         A     "DB123_MH_IO_Signals".MH[1].IN.MH_Stop;
         A     "DB123_MH_IO_Signals".MH[1].IN.MH_Manual_Mode;
   //    O
   //    UN    "DB005_RS<->Extern".FT_01.Daten_von_FT.Schaeumvorbereitung
         O     "DB123_MH_IO_Signals".MH[1].IN.MH_Auto_Mode;
         =     #Stop_MH;

         A     "DB123_MH_IO_Signals".MH[1].IN.MH_Status.shotactive_MH;
         AN    "DB614_MH_State".InertingMH[1].Inert_ON_OFF;
         A     "DB619_State_MPart".ShotMa[1].ShotData.PurgeMH_AfterShot;
         A     "DB614_MH_State".MH_Status[1].Switch_Service_ON_OFF;
         S     "DB614_MH_State".InertingMH[1].Start_Prepare_Purge_after_Shot;

         A     "DB614_MH_State".InertingMH[1].Start_Prepare_Purge_after_Shot;
         A     "DB619_State_MPart".Cycle[1].PulsShotend;
         A     "IPS_CP_MH01";
         S     "DB614_MH_State".InertingMH[1].Start_Purge_after_Shot;

         AN    "IPS_CP_MH01";
   //      U(
   //      U     "DB614_MH_State".InertingMH[1].Reserve41
   //      O     "DB614_MH_State".InertingMH[1].Inert_ON_OFF
   //      )
         A     "DB704_MH_Value".MH_Inerting[1].with_Purge;
         S     "DB614_MH_State".InertingMH[1].Enable_Purge;

         A     "IPS_CP_MH01";
         A     "DB614_MH_State".InertingMH[1].Enable_Purge;
         FP    "DB614_MH_State".InertingMH[1].Reserve40;
         S     "DB614_MH_State".InertingMH[1].Reserve42;

         A     "T_CP_forward_MH01";
         A     "DB614_MH_State".InertingMH[1].Enable_Purge;
         AN    "DB619_State_MPart".Cycle[1].running;
         S     "DB614_MH_State".InertingMH[1].Start_Purge_Manual;

         A     "DB614_MH_State".InertingMH[1].Start_Purge_Manual;
         AN    "DB619_State_MPart".Cycle[1].running;
         AN    "IPS_CP_MH01";
         S     "DB614_MH_State".InertingMH[1].HF_Start_Purge_Manual;
         R     "DB614_MH_State".InertingMH[1].Start_Purge_Manual;

         A(;
         A     "DB614_MH_State".InertingMH[1].HF_Start_Purge_Manual;
         O     "DB614_MH_State".InertingMH[1].Reserve42;
         );
         A     "IPS_CP_MH01";
         L     "DB704_MH_Value".MH_Inerting[1].Purge_time;
         JC    BLAS;

         A     "DB614_MH_State".InertingMH[1].Start_Purge_after_Shot;
         L     "DB704_MH_Value".MH_Inerting[1].Purge_after_Shot;
   BLAS: SE    "TM_Purge_after_Shot";
         A     "TM_Purge_after_Shot";
         FN    "DB614_MH_State".InertingMH[1].FN_Purge_after_shot_finished;
         R     "DB614_MH_State".InertingMH[1].HF_Start_Purge_Manual;
         R     "DB614_MH_State".InertingMH[1].Start_Prepare_Purge_after_Shot;
         R     "DB614_MH_State".InertingMH[1].Start_Purge_after_Shot;
         R     "DB614_MH_State".InertingMH[1].Enable_Purge;
         R     "DB614_MH_State".InertingMH[1].Reserve42;

         A     "TM_Purge_after_Shot";
         =     #Purge_Manual;

         A     #Purge_Manual;
         A     "DB614_MH_State".InertingMH[1].Reserve41;
         L     S5T#1S;
         SD    "TM_Reset_after_purge";
         A     "TM_Reset_after_purge";
         R     "DB704_MH_Value".MH_Inerting[1].with_purge_after_Shot;
         R     "DB614_MH_State".InertingMH[1].Enable_Purge;
         R     "DB614_MH_State".InertingMH[1].Reserve42;
         R     "DB614_MH_State".InertingMH[1].Reserve41;
         R     "DB614_MH_State".InertingMH[1].Start_Prepare_Purge_after_Shot;
         R     "DB614_MH_State".InertingMH[1].Start_Purge_after_Shot;

         L     0.0;
         T     "DB704_MH_Value".MH_Inerting[1].Reference_Value_Inert;

   //      CALL  "FC118_Enable_Inerting"
   //         Prg_Number     :=#InertPRG
   //         Ps_Number      :=1      //"DB619_State_MPart".ToolMa[1].PartShot
   //         ReferenceValue :="DB704_MH_Value".MH_Inerting[1].Reference_Value_Inert
   //         Inerting_OFF   :="DB614_MH_State".InertingMH[1].Inert_ON_OFF
   //         Shotwight      :=#Shotwight
END_REGION

REGION Network 2: MH01: Valve Nitrogen for Inerting
         SET;
         =     "DB704_MH_Value".MH_Inerting[1].with_Cycle_before_Inert_finished;

         CALL  "FC116_Inerting"
         ( IN_Enable                        := "DB619_State_MPart".Cycle[1].Release,
           IN_With_Inerting                 := "DB704_MH_Value".Mixinghead[1].WithInerting,
           IN_OP_Mode_Manual                := "DB123_MH_IO_Signals".MH[1].IN.MH_Manual_Mode,
           IN_OP_Mode_Wetshot               := 1,  //"DB614_MH_State".MH_Status[1].Switch_Service_ON_OFF
           IN_OP_Mode_Test                  := "DB619_State_MPart".Operationmode[1].Test,
           IN_Start                         := #Start_MH,
           IN_Stop                          := #Stop_MH,
           IN_T_Flushing                    := FALSE,
           IN_T_Purge_Air                   := #Purge_Manual,
           IN_Enable_pressurize_time        := "DB704_MH_Value".MH_Inerting[1].with_Cycle_before_Inert_finished,
           IN_AutoPurge_Air                 := FALSE,
           IN_Quitt_Fault                   := "DB009_Faults".Faults_Reset_FKT_M1,
           IN_Cycle_runs                    := FALSE,
           IN_MC_Activ                      := "DB614_MH_State".MH_Status[1].Switch_Service_ON_OFF,
           IN_PressurizeTimeRuns            := "DB619_State_MPart".Cycle[1].PressurizeTimeRuns,
           IN_Shotend                       := "DB619_State_MPart".Cycle[1].LastShotinToolFinished,
           IN_S_P_N2                        := "P_Nitrogen_Inerting_OK",
           IN_S_P_FlushingAgent             := TRUE,
           IN_MH_selected                   := "DB619_State_MPart".SWU[1].SWU_released."01",
           IN_Inert_MH                      := "DB704_MH_Value".MH_Inerting[1].with_inert_over_MH,
           IN_Inert_Lance                   := "DB704_MH_Value".MH_Inerting[1].with_inert_over_Lance,
           IN_IntervalCleaning              := "DB704_MH_Value".MH_Inerting[1].with_Interval_Purge,
           IN_Ctrl_Fault_On                 := TRUE,
           IN_Flowrate_N2_Actual            := "DB614_MH_State".InertingMH[1].Actual_Flow_N2_Visu,
           IN_Shotwight                     := #Shotwight,
           IN_Foam_Density                  := "DB704_MH_Value".MH_Inerting[1].Foam_density,
           IN_Leakage_value                 := "DB704_MH_Value".MH_Inerting[1].Leakage_Value,
           IN_DW_P_Build_Up_Before_Shot     := "DB700_Machine".Machine[1].PressureBuildUpTime,
           IN_DW_MaxInertTime               := "DB704_MH_Value".MH_Inerting[1].Max_Inerting_Time,
           IN_DW_Delay_Purge                := "DB704_MH_Value".MH_Inerting[1].Delay_Purge,
           IN_DW_Ready_time                 := "DB704_MH_Value".MH_Inerting[1].Ready_Time_after_Inert,
           IN_DW_Purge_time                 := "DB704_MH_Value".MH_Inerting[1].Purge_time,
           IN_DW_Delay_Plunger              := "DB704_MH_Value".MH_Inerting[1].Delay_Plunger,
           IN_DW_Delay_IntervalCleaning     := "DB704_MH_Value".MH_Inerting[1].Delay_Purge_Interval,
           IN_DW_PurgeTime_IntervalCleaning := "DB704_MH_Value".MH_Inerting[1].Purge_Time_interval,
           IN_DW_PauseTime_IntervalCleaning := "DB704_MH_Value".MH_Inerting[1].Pause_Time_interval,
           IN_DW_Duration_IntervalCleaning  := "DB704_MH_Value".MH_Inerting[1].Duration_Time_Interval,
           IN_Timer_Delay_Leakage           := "T_Leakage_Ctrl_N2",
           IN_Timer_hourly_tact             := "T_Leakage_Ctrl_Tact_N2",
           IN_Timer_Inerting                := "T_Inerting",
           IN_Timer_Ready                   := "T_Ready_for_Shot",
           IN_Timer_Delay_Purge             := "T_Delay_Purge",
           IN_Timer_Purge                   := "T_Purge",
           IN_Timer_Maximum_InertTime       := "T_Max_Inerting",
           IN_Timer_Delay_Plunger_N2        := "T_Delay_Plunger",
           IN_Timer_Delay_Tact              := "T_Delay_Purge_Tact",
           IN_Timer_PurgeTime_Tact          := "T_Purge_Tact",
           IN_Timer_PauseTime_Tact          := "T_Pause_Tact",
           IN_Timer_TotalTime_Tact          := "T_Total_Time_Purge",
           OUT_H_Inert                      := #dummy,
           OUT_H_Purge                      := #dummy,
           OUT_H_FlushingAgent              := #dummy,
           IO_DD_Inertfactor                := "DB704_MH_Value".MH_Inerting[1].Inerting_factor,
           IO_DD_StartOffset                := "DB704_MH_Value".MH_Inerting[1].Start_Offset,
           IO_DD_DF_N2_SetValue             := "DB614_MH_State".InertingMH[1].Computed_Value,
           IO_DD_DF_N2_Total                := "DB614_MH_State".InertingMH[1].Total_Flow_N2_Visu,
           IO_DD_DF_N2_Leakage              := "DB614_MH_State".InertingMH[1].Leakage_Total_Flow_N2_Visu,
           IO_MH_Logged_on                  := #dummy,
           IO_V_Piston                      := "V_Inert_Piston_MH1",
           IO_V_Inert                       := #Inerting,
           IO_V_Purge_Air                   := #Purge,
           IO_V_FlushingAgent               := #dummy,
           IO_Status                        := "DB614_MH_State".InertingMH[1],
           IO_Status_Faults                 := "DB824_Error_MH_CP".InertingBlowOut_MH[1],
           IO_NewFault                      := "DB009_Faults".Faultschanging_M1,
           IO_FaultLevel_1                  := "DB009_Faults".Faults_FKT_Grp_1_M1,
           IO_FaultLevel_2                  := "DB009_Faults".Faults_FKT_Grp_2_M1,
           IO_FaultLevel_3                  := "DB009_Faults".Faults_FKT_Grp_3_M1
         );

         A     #Purge;
         O     #Inerting;
         =     "V_Inert_MH1";
END_REGION
END_FUNCTION_BLOCK

FUNCTION_BLOCK "FB120_ProcanIO_RW"   // FB120, STL
TITLE = Transfer IO-Values from and to the ProCan-Moduls
{ S7_Optimized_Access := 'FALSE' }
AUTHOR : KT242
NAME : StPUCSPS
VERSION : 0.1
   VAR_TEMP
      Temp_ShotTimeAct : Real;
      dummy : Bool;
      Null : Word;
      ERROR_CODE : Int;
   END_VAR
BEGIN

REGION Network 1: Reset adresses od flow and MH
END_REGION

REGION Network 2: Read input values of procan modul
   //
         CALL  "FC120_read_ProCan";
END_REGION

REGION Network 3: PV Shot time
         L     0;
         T     #Temp_ShotTimeAct;

         AN    "DB619_State_MPart".SWU[1].Open_SWU_allone."01";
         JC    szm2;
         L     "DB123_MH_IO_Signals".MH[1].IN.Shottime;
         JU    szpv;
   szm2: AN    "DB619_State_MPart".SWU[1].Open_SWU_allone."02";
         JC    szm3;
         L     "DB123_MH_IO_Signals".MH[2].IN.Shottime;
         JU    szpv;
   szm3: AN    "DB619_State_MPart".SWU[1].Open_SWU_allone."03";
         JC    szm4;
         L     "DB123_MH_IO_Signals".MH[3].IN.Shottime;
         JU    szpv;
   szm4: AN    "DB619_State_MPart".SWU[1].Open_SWU_allone."04";
         JC    szm5;
         L     "DB123_MH_IO_Signals".MH[4].IN.Shottime;
         JU    szpv;
   szm5: AN    "DB619_State_MPart".SWU[1].Open_SWU_allone."05";
         JC    szm6;
         L     "DB123_MH_IO_Signals".MH[5].IN.Shottime;
         JU    szpv;
   szm6: AN    "DB619_State_MPart".SWU[1].Open_SWU_allone."06";
         JC    szm7;
         L     "DB123_MH_IO_Signals".MH[6].IN.Shottime;
         JU    szpv;
   szm7: AN    "DB619_State_MPart".SWU[1].Open_SWU_allone."07";
         JC    szm8;
         L     "DB123_MH_IO_Signals".MH[7].IN.Shottime;
         JU    szpv;
   szm8: AN    "DB619_State_MPart".SWU[1].Open_SWU_allone."08";
         JC    szm9;
         L     "DB123_MH_IO_Signals".MH[8].IN.Shottime;
         JU    szpv;
   szm9: AN    "DB619_State_MPart".SWU[1].Open_SWU_allone."09";
         JC    szm10;
         L     "DB123_MH_IO_Signals".MH[9].IN.Shottime;
         JU    szpv;
   szm10:AN    "DB619_State_MPart".SWU[1].Open_SWU_allone."10";
         JC    szm11;
         L     "DB123_MH_IO_Signals".MH[10].IN.Shottime;
         JU    szpv;
   szm11:AN    "DB619_State_MPart".SWU[1].Open_SWU_allone."11";
         JC    szm12;
         L     "DB123_MH_IO_Signals".MH[11].IN.Shottime;
         JU    szpv;
   szm12:AN    "DB619_State_MPart".SWU[1].Open_SWU_allone."12";
         JC    szm13;
         L     "DB123_MH_IO_Signals".MH[12].IN.Shottime;
         JU    szpv;
   szm13:JU    send;

   szpv: T     #Temp_ShotTimeAct;

         CALL  "FC920_PV_Calc_Act_Value"
         ( IN_Act_Value_read := TRUE,
           IN_Act_Value_ext  := TRUE,
           IN_Ext_Value      := #Temp_ShotTimeAct,
           IN_Read_Double    := TRUE,
           IN_FLT_Needful    := TRUE,
           IN_FLT_Reset      := "DB009_Faults".Faults_Reset_FKT_M1,
           IO_Any_ArrayPV    := "DB606_PV_Machine".Machine[1].ShotTime,
           IO_Fault_Sensor   := #dummy,
           IO_New_Fault      := #dummy,
           IO_FLT_Level_3    := #dummy
         );

   send: NOP   0;
END_REGION

REGION Network 4: Write output values of procan modul
   // Ein beschreiben der Module für die Mischköpfe ist nur bei LFI- Mischköpfen oder 
   // bei weiteren Mischköopfen bei dennen der Durchfluß eines Mediums am Mischkopf 
   // aufgenommen und geregelt wird (z.B. Faser) nötig.
   //
         CALL  "FC126_write_ProCan";
END_REGION
END_FUNCTION_BLOCK

FUNCTION_BLOCK "FB916_PV_LimitControl"   // FB916, STL
TITLE = Read prozess values and limit control of process values
{ S7_Optimized_Access := 'FALSE' }
AUTHOR : KT242
VERSION : 0.1
   VAR_TEMP
      DInt_dummy : DInt;
      FLT_quit_from_PLC : Bool;
      NewFault : Bool;
      ErrorLevel1 : Bool;
      ErrorLevel2 : Bool;
      ErrorLevel3 : Bool;
      TempStartTolTest : Bool;
      dummy : Bool;
      TempSwitchOffControl : Bool;
      CompForShotM1 : Array[1..16] of Bool;
      CompForShotM2 : Array[1..16] of Bool;
      PressureDiff : DInt;
      Temp_Con1MHConnected : Bool;
      Temp_Con2MHConnected : Bool;
      Temp_Con3MHConnected : Bool;
      Temp_Con4MHConnected : Bool;
      Temp_Con5MHConnected : Bool;
      Temp_Con6MHConnected : Bool;
      Temp_Con7MHConnected : Bool;
      Temp_Con8MHConnected : Bool;
   END_VAR
BEGIN

REGION Network 1: Actual pressure components at metering unit
         CALL  "FC_ActPressureMeteringUnit";
END_REGION

REGION Network 2: Actual values from mixinghead // temperatue and pressure
         CALL  "FC_ActValueMH";
END_REGION

REGION Network 3: Read tank temperatures -> FB101...
END_REGION

REGION Network 4: Limits of tank temperatures -> FB101...
END_REGION

REGION Network 5: Components for shot to local bits
         L;
         LAR1;
         L     "DB619_State_MPart".ShotMa[1].ShotData.Comp_at_Shot;
         CAW;
         T     LW[AR1, P#0.0];

         L;
         LAR1;
         L     "DB619_State_MPart".ShotMa[2].ShotData.Comp_at_Shot;
         CAW;
         T     LW[AR1, P#0.0];
END_REGION

REGION Network 6: Beim öffnen des MK die Überwachung um 500ms verzögern
         A     "DB619_State_MPart".Cycle[1].ShotRuns;
         L     s5t#500ms;
         SE    "TM_Delay_Limit_Control";
         A     "TM_Delay_Limit_Control";
         =     #TempSwitchOffControl;
END_REGION

REGION Network 7: Limits of flow pump component machine 1
         CALL  "FC_ToleranceValuesComponent"
         ( CompForShot      := #CompForShotM1,
           SwitchOffControl := #TempSwitchOffControl
         );
END_REGION

REGION Network 8: Limit foaming time
         A     "ShotStoppedM1";
         =     #TempStartTolTest;

         CALL  "FC916_PV_Limits"
         ( IN_Tolerance_Test     := #TempStartTolTest,
           IN_Reset_Fault        := "DB009_Faults".Faults_Reset_FKT_M1,
           IO_Any_ArrayPV        := "DB606_PV_Machine".Machine[1].ShotTime,
           IO_Fault_Warn_upperL  := "DB829_Error_Machine".Foaming_Time[1].Warning_limit_plus,
           IO_Fault_Warn_lowerL  := "DB829_Error_Machine".Foaming_Time[1].Warning_limit_minus,
           IO_Fault_Alarm_upperL := "DB829_Error_Machine".Foaming_Time[1].Alarm_limit_plus,
           IO_Fault_Alarm_lowerL := "DB829_Error_Machine".Foaming_Time[1].Alarm_limit_minus,
           IO_New_Fault          := "DB009_Faults".Faultschanging_M1,
           IO_Fault_Level_1      := "DB009_Faults".Faults_FKT_Grp_1_M1,
           IO_Fault_Level_2      := "DB009_Faults".Faults_FKT_Grp_2_M1,
           IO_Fault_Level_3      := "DB009_Faults".Faults_FKT_Grp_3_M1
         );
END_REGION

REGION Network 9: Sensor fault and warning and alarm limits Mixinghead Machine 1
         O     "DB614_MH_State".MH_Status[1].Switch_Testshot_A_ON_OFF;
         O     "DB614_MH_State".MH_Status[1].Switch_Testshot_B_ON_OFF;
         =     #dummy;

         CALL  "FC_ToleranceValuesMH"
         ( CompForShot      := #CompForShotM1,
           SwitchOffControl := #dummy  //FALSE
         );
   //---------
END_REGION

REGION Network 10: Read flow nitrogen
   //      CALL  "FC920_PV_Calc_Act_Value"
   //         IN_Act_Value_read :="DB704_MH_Value".Mixinghead[1].WithInerting
   //         IN_Act_Value_ext  :=FALSE
   //         IN_Ext_Value      :=#DInt_dummy
   //         IN_Read_Double    :=FALSE
   //         IN_FLT_Needful    :=TRUE
   //         IN_FLT_Reset      :="DB009_Faults".Faults_Reset_FKT_M1
   //         IO_Any_ArrayPV    :="DB604_PV_Mixinghead".Mixinghead[1].Inerting
   //         IO_Fault_Sensor   :="DB824_Error_MH_CP".InertingBlowOut_MH[1].Sensor_FLT_broken_wire
   //         IO_New_Fault      :="DB009_Faults".Faultschanging_M1
   //         IO_FLT_Level_3    :="DB009_Faults".Faults_FKT_Grp_3_M1

   //      L     "DB604_PV_Mixinghead".Mixinghead[1].Inerting.PV_ActV.Value
   //      T     "DB614_MH_State".InertingMH[1].Actual_Flow_N2
END_REGION
END_FUNCTION_BLOCK

FUNCTION_BLOCK "FB919_PV_SetValueFoaming"   // FB919, STL
TITLE = Set values flow component and pressure, temp. connected on MH
{ S7_Optimized_Access := 'FALSE' }
AUTHOR : KT242
VERSION : 0.1
   VAR_TEMP
      Temp_Shot_Time : DInt;
      Temp_Flow_C1 : DInt;
      Temp_Flow_C2 : DInt;
      Temp_Flow_C3 : DInt;
      Temp_Flow_C4 : DInt;
      Temp_OU_MR_C1 : DInt;
      Temp_OU_MR_C2 : DInt;
      Temp_OU_MR_C3 : DInt;
      Temp_OU_MR_C4 : DInt;
      Temp_IN_MR : DInt;
      dummyValue : DInt;
      DINT_dummy : DInt;
      MachineNo : Int;
      TempRetVal : Int;
      Temp_MHNumber_M1 : Int;
      Temp_MHNumber_M2 : Int;
      Temp_AmountComponent_M1 : Byte;
      Temp_AmountComponent_M2 : Byte;
      dummy : Bool;
   END_VAR
BEGIN

REGION Network 1
         L     0.0;
         AN    "DB619_State_MPart".Machine[1].Metering."01";
         AN    "DB619_State_MPart".Machine[1].Metering."02";
         JCN   Mxr0;

         T     "DB608_PV_Metering".Metering[1].MixingRatio.PV_ActV.Value;
         T     "DB608_PV_Metering".Metering[2].MixingRatio.PV_ActV.Value;
         T     "DB608_PV_Metering".Metering[3].MixingRatio.PV_ActV.Value;
         T     "DB608_PV_Metering".Metering[4].MixingRatio.PV_ActV.Value;
         T     "DB608_PV_Metering".Metering[5].MixingRatio.PV_ActV.Value;
         T     "DB608_PV_Metering".Metering[6].MixingRatio.PV_ActV.Value;
         T     "DB608_PV_Metering".Metering[7].MixingRatio.PV_ActV.Value;
         T     "DB608_PV_Metering".Metering[8].MixingRatio.PV_ActV.Value;

   Mxr0: NOP   0;
END_REGION

REGION Network 2
         L     0;
         T     #Temp_MHNumber_M1;
         T     #Temp_MHNumber_M2;
         T     #Temp_AmountComponent_M1;
         T     #Temp_AmountComponent_M2;
END_REGION

REGION Network 3: Select component at mixighead and flow of pump
   //---- Mixinghead 1 -----------------------------------------
         A(;
         O(;
         L     "DB619_State_MPart".ShotMa[1].ShotData.MH_No;
         L     1;
         <>I;
         A     "DB619_State_MPart".Cycle[1].running;
         );
         O(;
         AN    "DB619_State_MPart".SWU[1].Open_SWU."01";
         AN    "DB619_State_MPart".Cycle[1].running;
         );
         );
         A(;
         O(;
         L     "DB619_State_MPart".ShotMa[2].ShotData.MH_No;
         L     1;
         <>I;
         A     "DB619_State_MPart".Cycle[2].running;
         );
         O(;
         AN    "DB619_State_MPart".SWU[2].Open_SWU."01";
         AN    "DB619_State_MPart".Cycle[2].running;
         );
         );
         AN    "DB824_Error_MH_CP".MH_Control[1].FLTCompNotOnThisMH;
         JC    swu2;
   //---- Machine 1 MH 1 --------------------------------------
         L     "DB704_MH_Value".Mixinghead[1].MachineNumber;  // Example: If you have more than
         L     1;  // one machine you have to check
         ==D;  // whether the MH is connected to this machine
         JCN   M201;
   //-----
         L     1;
         T     #Temp_MHNumber_M1;
         L     "DB704_MH_Value".Mixinghead[1].AmountComponent;
         T     #Temp_AmountComponent_M1;
   //-----
         JU    swu2;
   //---- Machine 2 MH 1 ---------------------------------------
   M201: L     "DB704_MH_Value".Mixinghead[1].MachineNumber;  // Example: If you have more than
         L     2;  // one machine you have to check
         ==D;  // whether the MH is connected to this machine
         JCN   M301;
   //-----
         L     1;
         T     #Temp_MHNumber_M2;
         L     "DB704_MH_Value".Mixinghead[1].AmountComponent;
         T     #Temp_AmountComponent_M2;
   //-----
   M301: JU    swu2;
   //-----
   swu2: A(;
         O(;
         L     "DB619_State_MPart".ShotMa[1].ShotData.MH_No;
         L     2;
         <>I;
         A     "DB619_State_MPart".Cycle[1].running;
         );
         O(;
         AN    "DB619_State_MPart".SWU[1].Open_SWU."02";
         AN    "DB619_State_MPart".Cycle[1].running;
         );
         );
         A(;
         O(;
         L     "DB619_State_MPart".ShotMa[2].ShotData.MH_No;
         L     2;
         <>I;
         A     "DB619_State_MPart".Cycle[2].running;
         );
         O(;
         AN    "DB619_State_MPart".SWU[2].Open_SWU."02";
         AN    "DB619_State_MPart".Cycle[2].running;
         );
         );
         AN    "DB824_Error_MH_CP".MH_Control[2].FLTCompNotOnThisMH;
         JC    swu3;

   //---- Machine 1 MH 2 --------------------------------------
         L     "DB704_MH_Value".Mixinghead[2].MachineNumber;  // Example: If you have more than
         L     1;  // one machine you have to check
         ==D;  // whether the MH is connected to this machine
         JCN   M202;
   //-----
         L     2;
         T     #Temp_MHNumber_M1;
         L     "DB704_MH_Value".Mixinghead[2].AmountComponent;
         T     #Temp_AmountComponent_M1;
   //-----
         JU    swu3;
   //---- Machine 2 MH 2 ---------------------------------------
   M202: L     "DB704_MH_Value".Mixinghead[2].MachineNumber;  // Example: If you have more than
         L     2;  // one machine you have to check
         ==D;  // whether the MH is connected to this machine
         JCN   M302;
   //-----
         L     2;
         T     #Temp_MHNumber_M2;
         L     "DB704_MH_Value".Mixinghead[2].AmountComponent;
         T     #Temp_AmountComponent_M2;
   //-----
   M302: JU    swu3;

   //---- Mixinghead 3 -----------------------------------------
   swu3: A(;
         O(;
         L     "DB619_State_MPart".ShotMa[1].ShotData.MH_No;
         L     3;
         <>I;
         A     "DB619_State_MPart".Cycle[1].running;
         );
         O(;
         AN    "DB619_State_MPart".SWU[1].Open_SWU."03";
         AN    "DB619_State_MPart".Cycle[1].running;
         );
         );
         A(;
         O(;
         L     "DB619_State_MPart".ShotMa[2].ShotData.MH_No;
         L     3;
         <>I;
         A     "DB619_State_MPart".Cycle[2].running;
         );
         O(;
         AN    "DB619_State_MPart".SWU[2].Open_SWU."03";
         AN    "DB619_State_MPart".Cycle[2].running;
         );
         );
         AN    "DB824_Error_MH_CP".MH_Control[3].FLTCompNotOnThisMH;
         JC    swu4;
   //-----
         L     3;
         T     #Temp_MHNumber_M1;
         L     "DB704_MH_Value".Mixinghead[3].AmountComponent;
         T     #Temp_AmountComponent_M1;
   //-----

   //---- Mixinghead 4 -----------------------------------------
   swu4: A(;
         O(;
         L     "DB619_State_MPart".ShotMa[1].ShotData.MH_No;
         L     4;
         <>I;
         A     "DB619_State_MPart".Cycle[1].running;
         );
         O(;
         AN    "DB619_State_MPart".SWU[1].Open_SWU."04";
         AN    "DB619_State_MPart".Cycle[1].running;
         );
         );
         A(;
         O(;
         L     "DB619_State_MPart".ShotMa[2].ShotData.MH_No;
         L     4;
         <>I;
         A     "DB619_State_MPart".Cycle[2].running;
         );
         O(;
         AN    "DB619_State_MPart".SWU[2].Open_SWU."04";
         AN    "DB619_State_MPart".Cycle[2].running;
         );
         );
         AN    "DB824_Error_MH_CP".MH_Control[4].FLTCompNotOnThisMH;
         JC    swu5;

   //-----
         L     4;
         T     #Temp_MHNumber_M1;
         L     "DB704_MH_Value".Mixinghead[4].AmountComponent;
         T     #Temp_AmountComponent_M1;
         JU    swu5;
   //-----
   //---- Mixinghead 5 -----------------------------------------
   swu5: A(;
         O(;
         L     "DB619_State_MPart".ShotMa[1].ShotData.MH_No;
         L     5;
         <>I;
         A     "DB619_State_MPart".Cycle[1].running;
         );
         O(;
         AN    "DB619_State_MPart".SWU[1].Open_SWU."05";
         AN    "DB619_State_MPart".Cycle[1].running;
         );
         );
         A(;
         O(;
         L     "DB619_State_MPart".ShotMa[2].ShotData.MH_No;
         L     5;
         <>I;
         A     "DB619_State_MPart".Cycle[2].running;
         );
         O(;
         AN    "DB619_State_MPart".SWU[2].Open_SWU."05";
         AN    "DB619_State_MPart".Cycle[2].running;
         );
         );
         AN    "DB824_Error_MH_CP".MH_Control[5].FLTCompNotOnThisMH;
         JC    swu6;
   //-----
         L     5;
         T     #Temp_MHNumber_M1;
         L     "DB704_MH_Value".Mixinghead[5].AmountComponent;
         T     #Temp_AmountComponent_M1;
         JU    swu6;
   //-----
   //---- Mixinghead 6 -----------------------------------------
   swu6: A(;
         O(;
         L     "DB619_State_MPart".ShotMa[1].ShotData.MH_No;
         L     6;
         <>I;
         A     "DB619_State_MPart".Cycle[1].running;
         );
         O(;
         AN    "DB619_State_MPart".SWU[1].Open_SWU."06";
         AN    "DB619_State_MPart".Cycle[1].running;
         );
         );
         A(;
         O(;
         L     "DB619_State_MPart".ShotMa[2].ShotData.MH_No;
         L     6;
         <>I;
         A     "DB619_State_MPart".Cycle[2].running;
         );
         O(;
         AN    "DB619_State_MPart".SWU[2].Open_SWU."06";
         AN    "DB619_State_MPart".Cycle[2].running;
         );
         );
         AN    "DB824_Error_MH_CP".MH_Control[6].FLTCompNotOnThisMH;
         JC    swu7;
   //-----
         L     6;
         T     #Temp_MHNumber_M1;
         L     "DB704_MH_Value".Mixinghead[6].AmountComponent;
         T     #Temp_AmountComponent_M1;
         JU    swu7;
   //-----
   //---- Mixinghead 7 -----------------------------------------
   swu7: A(;
         O(;
         L     "DB619_State_MPart".ShotMa[1].ShotData.MH_No;
         L     7;
         <>I;
         A     "DB619_State_MPart".Cycle[1].running;
         );
         O(;
         AN    "DB619_State_MPart".SWU[1].Open_SWU."07";
         AN    "DB619_State_MPart".Cycle[1].running;
         );
         );
         A(;
         O(;
         L     "DB619_State_MPart".ShotMa[2].ShotData.MH_No;
         L     7;
         <>I;
         A     "DB619_State_MPart".Cycle[2].running;
         );
         O(;
         AN    "DB619_State_MPart".SWU[2].Open_SWU."07";
         AN    "DB619_State_MPart".Cycle[2].running;
         );
         );
         AN    "DB824_Error_MH_CP".MH_Control[7].FLTCompNotOnThisMH;
         JC    swu8;
   //-----
         L     7;
         T     #Temp_MHNumber_M1;
         L     "DB704_MH_Value".Mixinghead[7].AmountComponent;
         T     #Temp_AmountComponent_M1;
         JU    swu8;
   //-----
   //---- Mixinghead 8 -----------------------------------------
   swu8: A(;
         O(;
         L     "DB619_State_MPart".ShotMa[1].ShotData.MH_No;
         L     8;
         <>I;
         A     "DB619_State_MPart".Cycle[1].running;
         );
         O(;
         AN    "DB619_State_MPart".SWU[1].Open_SWU."08";
         AN    "DB619_State_MPart".Cycle[1].running;
         );
         );
         A(;
         O(;
         L     "DB619_State_MPart".ShotMa[2].ShotData.MH_No;
         L     8;
         <>I;
         A     "DB619_State_MPart".Cycle[2].running;
         );
         O(;
         AN    "DB619_State_MPart".SWU[2].Open_SWU."08";
         AN    "DB619_State_MPart".Cycle[2].running;
         );
         );
         AN    "DB824_Error_MH_CP".MH_Control[8].FLTCompNotOnThisMH;
         JC    swu9;
   //-----
         L     4;
         T     #Temp_MHNumber_M1;
         L     "DB704_MH_Value".Mixinghead[4].AmountComponent;
         T     #Temp_AmountComponent_M1;
         JU    swu5;
   //-----
   //-----
         L     8;
         T     #Temp_MHNumber_M1;
         L     "DB704_MH_Value".Mixinghead[8].AmountComponent;
         T     #Temp_AmountComponent_M1;
         JU    swu9;
   //-----
   //---- Mixinghead 9 -----------------------------------------
   swu9: A(;
         O(;
         L     "DB619_State_MPart".ShotMa[1].ShotData.MH_No;
         L     9;
         <>I;
         A     "DB619_State_MPart".Cycle[1].running;
         );
         O(;
         AN    "DB619_State_MPart".SWU[1].Open_SWU."09";
         AN    "DB619_State_MPart".Cycle[1].running;
         );
         );
         A(;
         O(;
         L     "DB619_State_MPart".ShotMa[2].ShotData.MH_No;
         L     9;
         <>I;
         A     "DB619_State_MPart".Cycle[2].running;
         );
         O(;
         AN    "DB619_State_MPart".SWU[2].Open_SWU."09";
         AN    "DB619_State_MPart".Cycle[2].running;
         );
         );
         AN    "DB824_Error_MH_CP".MH_Control[9].FLTCompNotOnThisMH;
         JC    swu10;
   //-----
         L     9;
         T     #Temp_MHNumber_M1;
         L     "DB704_MH_Value".Mixinghead[9].AmountComponent;
         T     #Temp_AmountComponent_M1;
         JU    swu10;
   //-----
   //---- Mixinghead 10 -----------------------------------------
   swu10:A(;
         O(;
         L     "DB619_State_MPart".ShotMa[1].ShotData.MH_No;
         L     10;
         <>I;
         A     "DB619_State_MPart".Cycle[1].running;
         );
         O(;
         AN    "DB619_State_MPart".SWU[1].Open_SWU."10";
         AN    "DB619_State_MPart".Cycle[1].running;
         );
         );
         A(;
         O(;
         L     "DB619_State_MPart".ShotMa[2].ShotData.MH_No;
         L     10;
         <>I;
         A     "DB619_State_MPart".Cycle[2].running;
         );
         O(;
         AN    "DB619_State_MPart".SWU[2].Open_SWU."10";
         AN    "DB619_State_MPart".Cycle[2].running;
         );
         );
         AN    "DB824_Error_MH_CP".MH_Control[10].FLTCompNotOnThisMH;
         JC    swu11;
   //-----
         L     10;
         T     #Temp_MHNumber_M1;
         L     "DB704_MH_Value".Mixinghead[10].AmountComponent;
         T     #Temp_AmountComponent_M1;
         JU    swu11;
   //-----
   //---- Mixinghead 11 -----------------------------------------
   swu11:NOP   0;
END_REGION

REGION Network 4
         L     #Temp_MHNumber_M1;
         L     0;
         <>I;
         JC    GetValue;
   // When No MH is activ set Mixing ratio to 100% and Exit
   //      L     100.0
   //      T     "DB608_PV_Metering".Metering[1].MixingRatio.PV_ActV.Value
   //      T     "DB608_PV_Metering".Metering[2].MixingRatio.PV_ActV.Value
   //      T     "DB608_PV_Metering".Metering[3].MixingRatio.PV_ActV.Value
   //      T     "DB608_PV_Metering".Metering[4].MixingRatio.PV_ActV.Value
   //      T     "DB608_PV_Metering".Metering[5].MixingRatio.PV_ActV.Value
   //      T     "DB608_PV_Metering".Metering[6].MixingRatio.PV_ActV.Value
         BEU;
   GetValue:NOP   0;
   //-----
         CALL  "FC1156_FlowPressMH_Instance"
         ( IN_MachineNo            := 1,
           IN_MixingHeadNo         := #Temp_MHNumber_M1,
           IN_AmountMHConnections  := #Temp_AmountComponent_M1,
           IN_Cycle                := "DB619_State_MPart".Cycle[1].running,
           IN_ReducedRecirculation := "DB619_State_MPart".Recirculation[1].Reduced,
           IN_LPRecirculation      := "DB619_State_MPart".Recirculation[1].Lowpressure,
           IN_HPRecirculation      := "DB619_State_MPart".Recirculation[1].Highpressure,
           IN_PauseTime            := "DB619_State_MPart".Recirculation[1].Pausetime,
           IN_Reset_Fault          := "DB009_Faults".HF_Faults_Quit,
           IO_FaultWrongAssignment := "DB829_Error_Machine".PouringCycle[1].FLT_CompAllocation,
           IO_Fault_Level_1        := "DB009_Faults".Faults_FKT_Grp_1_M1,
           IO_New_Fault            := "DB009_Faults".Faultschanging_M1
         );
   //-----
END_REGION
END_FUNCTION_BLOCK

FUNCTION_BLOCK "FB920_ShotResult"   // FB920, STL
TITLE = Act.value mixing head temp.; shot results;
{ S7_Optimized_Access := 'FALSE' }
VERSION : 0.1
   VAR_TEMP
      DInt_dummy : DInt;
      CompUsedForShot : Array[1..16] of Bool;
      "Return" : Int;
      dummy : Bool;
   END_VAR
BEGIN

REGION Network 1
   // Copy Control bits for module to local area
         L;
         LAR1;
         L     "DB619_State_MPart".ShotMa[1].ShotData.Comp_at_Shot;
         CAW;
         T     LW[AR1, P#0.0];
   //-----
         A     "M_ShotActive";  // "DB610_State_MPart".Cycle_Ma[1].ShotRuns
         JCN   f1;

         CALL  "ShotData_01"
         ( CompForShot := #CompUsedForShot
         );
   //-----
   f1:   NOP   0;
   //-----
END_REGION

REGION Network 2: Temperature component tank machine 1
   // Tank temperatures of machine 1
         AN    "DB619_State_MPart".Cycle[1].ShotRuns;
         JC    TT1e;
   // Inerting

         L     "DB619_State_MPart".ActMHInerting[1].Total_Flow_N2_Visu;
         T     "DB919_ShotResultMach".ShotResult_Ma[1].General.NitrogenValue_Inerting;
   //
         L     "DB602_PV_Tank".Tank[1].Temp.PV_ActV.Value;
         T     "DB919_ShotResultMach".ShotResult_Ma[1].Component.Comp[1].Temperature;
         L     "DB602_PV_Tank".Tank[2].Temp.PV_ActV.Value;
         T     "DB919_ShotResultMach".ShotResult_Ma[1].Component.Comp[2].Temperature;
         L     "DB602_PV_Tank".Tank[3].Temp.PV_ActV.Value;
         T     "DB919_ShotResultMach".ShotResult_Ma[1].Component.Comp[3].Temperature;
         L     "DB602_PV_Tank".Tank[4].Temp.PV_ActV.Value;
         T     "DB919_ShotResultMach".ShotResult_Ma[1].Component.Comp[4].Temperature;
         L     "DB602_PV_Tank".Tank[5].Temp.PV_ActV.Value;
         T     "DB919_ShotResultMach".ShotResult_Ma[1].Component.Comp[5].Temperature;
         L     "DB602_PV_Tank".Tank[6].Temp.PV_ActV.Value;
         T     "DB919_ShotResultMach".ShotResult_Ma[1].Component.Comp[6].Temperature;

   TT1e: NOP   0;
END_REGION

REGION Network 3: Shot results machine 1 general values and componet values
         A     "DB619_State_MPart".Cycle[1].ShotRuns;
         FP    "FHM_ShotRunsMH1";
         JCN   M014;

         ON    "DB619_State_MPart".Operationmode[1].Operation;
         O     "DB619_State_MPart".ShotMa[1].ShotData.ShotDisabled;
         S     "DB919_ShotResultMach".ShotResult_Ma[1].General.ServiceShot;

         L     "DB619_State_MPart".ToolMa[1].StationNo;
         T     "DB919_ShotResultMach".ShotResult_Ma[1].General.StationNo;

         L     "DB619_State_MPart".ShotMa[1].ShotData.MH_No;
         T     "DB919_ShotResultMach".ShotResult_Ma[1].General.MH_No;

         L     "DB619_State_MPart".ToolMa[1].ToolNo;
         T     "DB919_ShotResultMach".ShotResult_Ma[1].General.ToolNo;

         L     "DB619_State_MPart".ShotMa[1].ShotData.PartCounter;
         T     "DB919_ShotResultMach".ShotResult_Ma[1].General.PartID;

         L     1;
         T     "DB919_ShotResultMach".ShotResult_Ma[1].General.Machine_No;

         L     "CompAtShot";
         T     "DB919_ShotResultMach".ShotResult_Ma[1].General.MH_CompAlloc;

         AN    "DB619_State_MPart".Cycle[1].ShotRuns;
         JC    M014;

         L     "ShotNoNextMa1";  //  -> FB1930 GetToolShotValues
         T     "DB919_ShotResultMach".ShotResult_Ma[1].General.ShotNo;

         CALL  BLKMOV
         ( SRCBLK  := "DB619_State_MPart".ActMHComponent[1]."Name"[1],
           RET_VAL := #"Return",
           DSTBLK  := "DB919_ShotResultMach".ShotResult_Ma[1].Component.Comp[1]."Name"
         );
         CALL  BLKMOV
         ( SRCBLK  := "DB619_State_MPart".ActMHComponent[1]."Name"[2],
           RET_VAL := #"Return",
           DSTBLK  := "DB919_ShotResultMach".ShotResult_Ma[1].Component.Comp[2]."Name"
         );
         CALL  BLKMOV
         ( SRCBLK  := "DB619_State_MPart".ActMHComponent[1]."Name"[3],
           RET_VAL := #"Return",
           DSTBLK  := "DB919_ShotResultMach".ShotResult_Ma[1].Component.Comp[3]."Name"
         );
         CALL  BLKMOV
         ( SRCBLK  := "DB619_State_MPart".ActMHComponent[1]."Name"[4],
           RET_VAL := #"Return",
           DSTBLK  := "DB919_ShotResultMach".ShotResult_Ma[1].Component.Comp[4]."Name"
         );
         CALL  BLKMOV
         ( SRCBLK  := "DB619_State_MPart".ActMHComponent[1]."Name"[5],
           RET_VAL := #"Return",
           DSTBLK  := "DB919_ShotResultMach".ShotResult_Ma[1].Component.Comp[5]."Name"
         );
         CALL  BLKMOV
         ( SRCBLK  := "DB619_State_MPart".ActMHComponent[1]."Name"[6],
           RET_VAL := #"Return",
           DSTBLK  := "DB919_ShotResultMach".ShotResult_Ma[1].Component.Comp[6]."Name"
         );


   M014: A     "DB619_State_MPart".Cycle[1].ShotRuns;
         FN    "NoShotActiveM1";  // No shot active
         S     "ShotStoppedM1";  // Shot stopped
         AN    "NoShotActiveM1";
         JC    con1;

   //-----------------------------------------------------------------------------------
   //    Pressure mixinghead connection -> component at MH
   //-----------------------------------------------------------------------------------
         AN    "DB919_ShotResultMach".ShotResult_Ma[1].Component.Comp[1].ComponentActive;
         O     "DB614_MH_State".MH_Status[1].Switch_Testshot_B_ON_OFF;
         L     0.0;
         JC    NoPressureMHC1;
         L     "DB619_State_MPart".ActMHPressureMa[1].Comp[1];
   NoPressureMHC1:NOP   0;
         T     "DB919_ShotResultMach".ShotResult_Ma[1].Component.Comp[1].PressureMH;

         AN    "DB919_ShotResultMach".ShotResult_Ma[1].Component.Comp[2].ComponentActive;
         O     "DB614_MH_State".MH_Status[1].Switch_Testshot_A_ON_OFF;
         L     0.0;
         JC    NoPressureMHC2;
         L     "DB619_State_MPart".ActMHPressureMa[1].Comp[2];
   NoPressureMHC2:NOP   0;
         T     "DB919_ShotResultMach".ShotResult_Ma[1].Component.Comp[2].PressureMH;

         AN    "DB919_ShotResultMach".ShotResult_Ma[1].Component.Comp[3].ComponentActive;
         L     0.0;
         JC    NoPressureMHC3;
         L     "DB619_State_MPart".ActMHPressureMa[1].Comp[3];
   NoPressureMHC3:NOP   0;
         T     "DB919_ShotResultMach".ShotResult_Ma[1].Component.Comp[3].PressureMH;

         AN    "DB919_ShotResultMach".ShotResult_Ma[1].Component.Comp[4].ComponentActive;
         L     0.0;
         JC    NoPressureMHC4;
         L     "DB619_State_MPart".ActMHPressureMa[1].Comp[4];
   NoPressureMHC4:NOP   0;
         T     "DB919_ShotResultMach".ShotResult_Ma[1].Component.Comp[4].PressureMH;

         AN    "DB919_ShotResultMach".ShotResult_Ma[1].Component.Comp[5].ComponentActive;
         L     0.0;
         JC    NoPressureMHC5;
         L     "DB619_State_MPart".ActMHPressureMa[1].Comp[5];
   NoPressureMHC5:NOP   0;
         T     "DB919_ShotResultMach".ShotResult_Ma[1].Component.Comp[5].PressureMH;

         AN    "DB919_ShotResultMach".ShotResult_Ma[1].Component.Comp[6].ComponentActive;
         L     0.0;
         JC    NoPressureMHC6;
         L     "DB619_State_MPart".ActMHPressureMa[1].Comp[6];
   NoPressureMHC6:NOP   0;
         T     "DB919_ShotResultMach".ShotResult_Ma[1].Component.Comp[6].PressureMH;

   //-----------------------------------------------------------------------------------
   //    Pressure metering units 1 - 6
   //-----------------------------------------------------------------------------------
         L     "DB608_PV_Metering".Metering[1].Pressure.PV_ActV.Value;
         T     "DB919_ShotResultMach".ShotResult_Ma[1].Component.Comp[1].Pressure;
         L     "DB608_PV_Metering".Metering[2].Pressure.PV_ActV.Value;
         T     "DB919_ShotResultMach".ShotResult_Ma[1].Component.Comp[2].Pressure;
         L     "DB608_PV_Metering".Metering[3].Pressure.PV_ActV.Value;
         T     "DB919_ShotResultMach".ShotResult_Ma[1].Component.Comp[3].Pressure;
         L     "DB608_PV_Metering".Metering[4].Pressure.PV_ActV.Value;
         T     "DB919_ShotResultMach".ShotResult_Ma[1].Component.Comp[4].Pressure;
         L     "DB608_PV_Metering".Metering[5].Pressure.PV_ActV.Value;
         T     "DB919_ShotResultMach".ShotResult_Ma[1].Component.Comp[5].Pressure;
         L     "DB608_PV_Metering".Metering[6].Pressure.PV_ActV.Value;
         T     "DB919_ShotResultMach".ShotResult_Ma[1].Component.Comp[6].Pressure;
   // Set Values
         L     "DB608_PV_Metering".Metering[1].Pressure.PV_SetV.Value;
         T     "DB919_ShotResultMach".ShotResult_Ma[1].Component.Comp[1].Pressure_Set;
         L     "DB608_PV_Metering".Metering[2].Pressure.PV_SetV.Value;
         T     "DB919_ShotResultMach".ShotResult_Ma[1].Component.Comp[2].Pressure_Set;
         L     "DB608_PV_Metering".Metering[3].Pressure.PV_SetV.Value;
         T     "DB919_ShotResultMach".ShotResult_Ma[1].Component.Comp[3].Pressure_Set;
         L     "DB608_PV_Metering".Metering[4].Pressure.PV_SetV.Value;
         T     "DB919_ShotResultMach".ShotResult_Ma[1].Component.Comp[4].Pressure_Set;
         L     "DB608_PV_Metering".Metering[5].Pressure.PV_SetV.Value;
         T     "DB919_ShotResultMach".ShotResult_Ma[1].Component.Comp[5].Pressure_Set;
         L     "DB608_PV_Metering".Metering[6].Pressure.PV_SetV.Value;
         T     "DB919_ShotResultMach".ShotResult_Ma[1].Component.Comp[6].Pressure_Set;
   //-----------------------------------------------------------------------------------
   //    Flow - Set Values
   //-----------------------------------------------------------------------------------
         L     "DB608_PV_Metering".Metering[1].Flow.PV_SetV.Value;
         T     "DB919_ShotResultMach".ShotResult_Ma[1].Component.Comp[1].Flow_Set;
         L     "DB608_PV_Metering".Metering[2].Flow.PV_SetV.Value;
         T     "DB919_ShotResultMach".ShotResult_Ma[1].Component.Comp[2].Flow_Set;
         L     "DB608_PV_Metering".Metering[3].Flow.PV_SetV.Value;
         T     "DB919_ShotResultMach".ShotResult_Ma[1].Component.Comp[3].Flow_Set;
         L     "DB608_PV_Metering".Metering[4].Flow.PV_SetV.Value;
         T     "DB919_ShotResultMach".ShotResult_Ma[1].Component.Comp[4].Flow_Set;
         L     "DB608_PV_Metering".Metering[5].Flow.PV_SetV.Value;
         T     "DB919_ShotResultMach".ShotResult_Ma[1].Component.Comp[5].Flow_Set;
         L     "DB608_PV_Metering".Metering[6].Flow.PV_SetV.Value;
         T     "DB919_ShotResultMach".ShotResult_Ma[1].Component.Comp[6].Flow_Set;
   //-----------------------------------------------------------------------------------
   //    Temperature mixinghead connection -> component at MH
   //-----------------------------------------------------------------------------------
         AN    "DB919_ShotResultMach".ShotResult_Ma[1].Component.Comp[1].ComponentActive;
         O     "DB614_MH_State".MH_Status[1].Switch_Testshot_B_ON_OFF;
         L     0.0;
         JC    NoTempMHC1;
         L     "DB619_State_MPart".ActMHTemperatureMa[1].Comp[1];
   NoTempMHC1:NOP   0;
         T     "DB919_ShotResultMach".ShotResult_Ma[1].Component.Comp[1].TemperatureMH;

         AN    "DB919_ShotResultMach".ShotResult_Ma[1].Component.Comp[2].ComponentActive;
         O     "DB614_MH_State".MH_Status[1].Switch_Testshot_A_ON_OFF;
         L     0.0;
         JC    NoTempMHC2;
         L     "DB619_State_MPart".ActMHTemperatureMa[1].Comp[2];
   NoTempMHC2:NOP   0;
         T     "DB919_ShotResultMach".ShotResult_Ma[1].Component.Comp[2].TemperatureMH;

         AN    "DB919_ShotResultMach".ShotResult_Ma[1].Component.Comp[3].ComponentActive;
         L     0.0;
         JC    NoTempMHC3;
         L     "DB619_State_MPart".ActMHTemperatureMa[1].Comp[3];
   NoTempMHC3:NOP   0;
         T     "DB919_ShotResultMach".ShotResult_Ma[1].Component.Comp[3].TemperatureMH;

         AN    "DB919_ShotResultMach".ShotResult_Ma[1].Component.Comp[4].ComponentActive;
         L     0.0;
         JC    NoTempMHC4;
         L     "DB619_State_MPart".ActMHTemperatureMa[1].Comp[4];
   NoTempMHC4:NOP   0;
         T     "DB919_ShotResultMach".ShotResult_Ma[1].Component.Comp[4].TemperatureMH;

         AN    "DB919_ShotResultMach".ShotResult_Ma[1].Component.Comp[5].ComponentActive;
         L     0.0;
         JC    NoTempMHC5;
         L     "DB619_State_MPart".ActMHTemperatureMa[1].Comp[5];
   NoTempMHC5:NOP   0;
         T     "DB919_ShotResultMach".ShotResult_Ma[1].Component.Comp[5].TemperatureMH;

         AN    "DB919_ShotResultMach".ShotResult_Ma[1].Component.Comp[6].ComponentActive;
         L     0.0;
         JC    NoTempMHC6;
         L     "DB619_State_MPart".ActMHTemperatureMa[1].Comp[6];
   NoTempMHC6:NOP   0;
         T     "DB919_ShotResultMach".ShotResult_Ma[1].Component.Comp[6].TemperatureMH;

   con1: A     "CalcShotValuesMa1";  // Shot values detected after shot
         A     "ShotStoppedM1";  // Shot stopped
         JCN   SEM1;
         S     "DB918_ShotResultlast10".NewData;
         R     "CalcShotValuesMa1";
         R     "ShotStoppedM1";

         CALL  RD_SYS_T
         ( RET_VAL := #"Return",
           OUT     := "DB919_ShotResultMach".ShotResult_Ma[1].General.DateTime
         );

   //---------------------------------------------------------------------------------------
   //    Calculate part weight
   //---------------------------------------------------------------------------------------
         L     0.0;
         AN    "DB919_ShotResultMach".ShotResult_Ma[1].Component.Comp[1].ComponentActive;
         O     "DB614_MH_State".MH_Status[1].Switch_Testshot_B_ON_OFF;
         JC    NoConsumptionC1;
         L     "DB919_ShotResultMach".ShotResult_Ma[1].Component.Comp[1].MaterialConsumption;
         +R;
   NoConsumptionC1:NOP   0;
         AN    "DB919_ShotResultMach".ShotResult_Ma[1].Component.Comp[2].ComponentActive;
         O     "DB614_MH_State".MH_Status[1].Switch_Testshot_A_ON_OFF;
         JC    NoConsumptionC2;
         L     "DB919_ShotResultMach".ShotResult_Ma[1].Component.Comp[2].MaterialConsumption;
         +R;
   NoConsumptionC2:NOP   0;
         AN    "DB919_ShotResultMach".ShotResult_Ma[1].Component.Comp[3].ComponentActive;
         JC    NoConsumptionC3;
         L     "DB919_ShotResultMach".ShotResult_Ma[1].Component.Comp[3].MaterialConsumption;
         +R;
   NoConsumptionC3:NOP   0;
         AN    "DB919_ShotResultMach".ShotResult_Ma[1].Component.Comp[4].ComponentActive;
         JC    NoConsumptionC4;
         L     "DB919_ShotResultMach".ShotResult_Ma[1].Component.Comp[4].MaterialConsumption;
         +R;
   NoConsumptionC4:NOP   0;
         AN    "DB919_ShotResultMach".ShotResult_Ma[1].Component.Comp[5].ComponentActive;
         JC    NoConsumptionC5;
         L     "DB919_ShotResultMach".ShotResult_Ma[1].Component.Comp[5].MaterialConsumption;
         +R;
   NoConsumptionC5:NOP   0;
         AN    "DB919_ShotResultMach".ShotResult_Ma[1].Component.Comp[6].ComponentActive;
         JC    NoConsumptionC6;
         L     "DB919_ShotResultMach".ShotResult_Ma[1].Component.Comp[6].MaterialConsumption;
         +R;
   NoConsumptionC6:NOP   0;
         T     "DB919_ShotResultMach".ShotResult_Ma[1].General.PartWeight;

         L     0.0;
         A     "DB919_ShotResultMach".ShotResult_Ma[1].General.ServiceShot;
         JC    NoCorrValue;
         L     "DB704_MH_Value".Mixinghead[1].Corrvalue;  // Verzögerung des Steuerkolbens
   NoCorrValue:NOP   0;
         L     "DB606_PV_Machine".Machine[1].ShotTime.PV_ActV.Value;  // Korrigiere Zeit um eingestellte
         +R;
         T     "DB919_ShotResultMach".ShotResult_Ma[1].General.FoamingTime;

         L     "DB123_MH_IO_Signals".MH[1].IN.MH_Opentime;
         T     "DB919_ShotResultMach".ShotResult_Ma[1].General.MH_OpeningTime;

         L     "DB123_MH_IO_Signals".MH[1].IN.MH_Closingtime;
         T     "DB919_ShotResultMach".ShotResult_Ma[1].General.MH_CloseingTime;

         L     "DB919_ShotResultMach".ShotResult_Ma[1].General.ShotNo;
         L     1;
         <>I;
         JC    ntm1;

         CALL  RD_SYS_T
         ( RET_VAL := #"Return",
           OUT     := "DB919_ShotResultMach".ShotResult_Ma[1].General.ToolStartTime
         );

   ntm1: NOP   0;

   //------------------------------------------------------------------------------
   // Copy shotresult to shotbuffer finished -> VISU can read values
   //------------------------------------------------------------------------------
         AN    "DB919_ShotResultMach".ShotResult_Ma[1].General.ServiceShot;
         S     "BufferShotResultM1";

         SET;
         R     "DB919_ShotResultMach".ShotResult_Ma[1].General.ServiceShot;

         SET;  /// TEST
         S     "M_NewShotDataToMC";  // For traceability

   SEM1: NOP   0;

         A     "BufferShotResultM1";
         FP    "FP_BufferShotResultM1";
         JCN   m1;